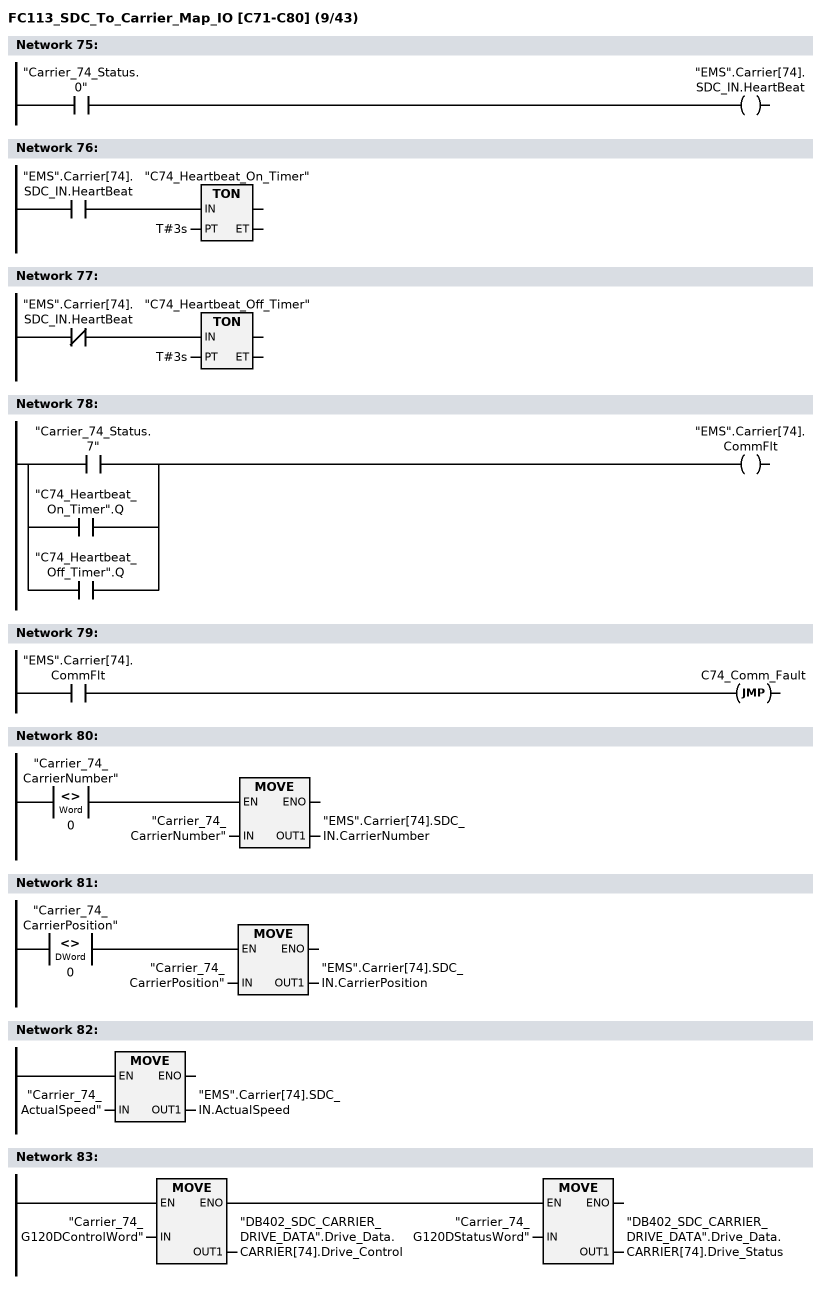
   RUNG wire#powerrail
      Contact( "Carrier_74_Status.0" )
      Coil( "EMS".Carrier[74].SDC_IN.HeartBeat )
   END_RUNG
   // the same network as SCL:
   "EMS".Carrier[74].SDC_IN.HeartBeat := "Carrier_74_Status.0";
END_REGION

REGION Network 76
   "C74_Heartbeat_On_Timer".TON(IN := "EMS".Carrier[74].SDC_IN.HeartBeat, PT := T#3s);
END_REGION

REGION Network 77
   "C74_Heartbeat_Off_Timer".TON(IN := NOT "EMS".Carrier[74].SDC_IN.HeartBeat, PT := T#3s);
END_REGION

REGION Network 78
   RUNG wire#powerrail
      Contact( "Carrier_74_Status.7" )
      wire#w1
      Coil( "EMS".Carrier[74].CommFlt )
   END_RUNG
   RUNG wire#powerrail
      Contact( "C74_Heartbeat_On_Timer".Q )
   END_RUNG wire#w1
   RUNG wire#powerrail
      Contact( "C74_Heartbeat_Off_Timer".Q )
   END_RUNG wire#w1
   // the same network as SCL:
   "EMS".Carrier[74].CommFlt := "Carrier_74_Status.7" OR "C74_Heartbeat_On_Timer".Q OR "C74_Heartbeat_Off_Timer".Q;
END_REGION

REGION Network 79
   RUNG wire#powerrail
      Contact( "EMS".Carrier[74].CommFlt )
      JumpCoil( C74_Comm_Fault )
   END_RUNG
   // the same network as SCL:
   IF "EMS".Carrier[74].CommFlt THEN GOTO C74_Comm_Fault; END_IF;
END_REGION

REGION Network 80
   RUNG wire#powerrail
      { S7_Templates := "SrcType := Word" } NE_Contact(in1 := "Carrier_74_CarrierNumber", in2 := 0)
      Move(in := "Carrier_74_CarrierNumber", out1 => "EMS".Carrier[74].SDC_IN.CarrierNumber)
   END_RUNG
   // the same network as SCL:
   IF "Carrier_74_CarrierNumber" <> 0 THEN
       "EMS".Carrier[74].SDC_IN.CarrierNumber := "Carrier_74_CarrierNumber";
   END_IF;
END_REGION

REGION Network 81
   RUNG wire#powerrail
      { S7_Templates := "SrcType := DWord" } NE_Contact(in1 := "Carrier_74_CarrierPosition", in2 := 0)
      Move(in := "Carrier_74_CarrierPosition", out1 => "EMS".Carrier[74].SDC_IN.CarrierPosition)
   END_RUNG
   // the same network as SCL:
   IF "Carrier_74_CarrierPosition" <> 0 THEN
       "EMS".Carrier[74].SDC_IN.CarrierPosition := "Carrier_74_CarrierPosition";
   END_IF;
END_REGION

REGION Network 82
   RUNG wire#powerrail
      Move(in := "Carrier_74_ActualSpeed", out1 => "EMS".Carrier[74].SDC_IN.ActualSpeed)
   END_RUNG
   // the same network as SCL:
   "EMS".Carrier[74].SDC_IN.ActualSpeed := "Carrier_74_ActualSpeed";
END_REGION

REGION Network 83
   RUNG wire#powerrail
      Move(in := "Carrier_74_G120DControlWord", out1 => "DB402_SDC_CARRIER_DRIVE_DATA".Drive_Data.CARRIER[74].Drive_Control)
      Move(in := "Carrier_74_G120DStatusWord", out1 => "DB402_SDC_CARRIER_DRIVE_DATA".Drive_Data.CARRIER[74].Drive_Status)
   END_RUNG
   // the same network as SCL:
   "DB402_SDC_CARRIER_DRIVE_DATA".Drive_Data.CARRIER[74].Drive_Control := "Carrier_74_G120DControlWord";
   "DB402_SDC_CARRIER_DRIVE_DATA".Drive_Data.CARRIER[74].Drive_Status := "Carrier_74_G120DStatusWord";
END_REGION

REGION Network 84
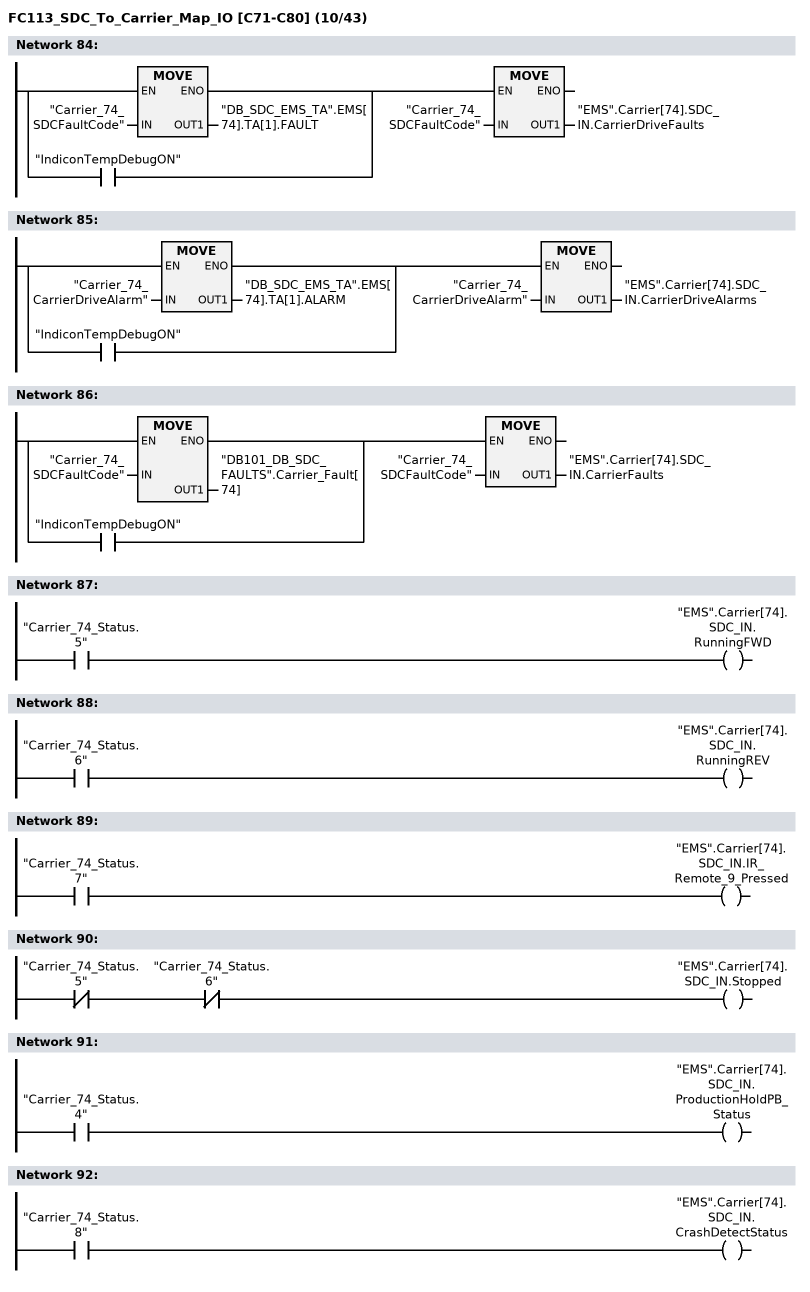
   RUNG wire#powerrail
      Move(in := "Carrier_74_SDCFaultCode", out1 => "DB_SDC_EMS_TA".EMS[74].TA[1].FAULT)
      wire#w1
      Move(in := "Carrier_74_SDCFaultCode", out1 => "EMS".Carrier[74].SDC_IN.CarrierDriveFaults)
   END_RUNG
   RUNG wire#powerrail
      Contact( "IndiconTempDebugON" )
   END_RUNG wire#w1
   // the same network as SCL:
   "DB_SDC_EMS_TA".EMS[74].TA[1].FAULT := "Carrier_74_SDCFaultCode";
   IF TRUE OR "IndiconTempDebugON" THEN
       "EMS".Carrier[74].SDC_IN.CarrierDriveFaults := "Carrier_74_SDCFaultCode";
   END_IF;
END_REGION

REGION Network 85
   RUNG wire#powerrail
      Move(in := "Carrier_74_CarrierDriveAlarm", out1 => "DB_SDC_EMS_TA".EMS[74].TA[1].ALARM)
      wire#w1
      Move(in := "Carrier_74_CarrierDriveAlarm", out1 => "EMS".Carrier[74].SDC_IN.CarrierDriveAlarms)
   END_RUNG
   RUNG wire#powerrail
      Contact( "IndiconTempDebugON" )
   END_RUNG wire#w1
   // the same network as SCL:
   "DB_SDC_EMS_TA".EMS[74].TA[1].ALARM := "Carrier_74_CarrierDriveAlarm";
   IF TRUE OR "IndiconTempDebugON" THEN
       "EMS".Carrier[74].SDC_IN.CarrierDriveAlarms := "Carrier_74_CarrierDriveAlarm";
   END_IF;
END_REGION

REGION Network 86
   RUNG wire#powerrail
      Move(in := "Carrier_74_SDCFaultCode", out1 => "DB101_DB_SDC_FAULTS".Carrier_Fault[74])
      wire#w1
      Move(in := "Carrier_74_SDCFaultCode", out1 => "EMS".Carrier[74].SDC_IN.CarrierFaults)
   END_RUNG
   RUNG wire#powerrail
      Contact( "IndiconTempDebugON" )
   END_RUNG wire#w1
   // the same network as SCL:
   "DB101_DB_SDC_FAULTS".Carrier_Fault[74] := "Carrier_74_SDCFaultCode";
   IF TRUE OR "IndiconTempDebugON" THEN
       "EMS".Carrier[74].SDC_IN.CarrierFaults := "Carrier_74_SDCFaultCode";
   END_IF;
END_REGION

REGION Network 87
   RUNG wire#powerrail
      Contact( "Carrier_74_Status.5" )
      Coil( "EMS".Carrier[74].SDC_IN.RunningFWD )
   END_RUNG
   // the same network as SCL:
   "EMS".Carrier[74].SDC_IN.RunningFWD := "Carrier_74_Status.5";
END_REGION

REGION Network 88
   RUNG wire#powerrail
      Contact( "Carrier_74_Status.6" )
      Coil( "EMS".Carrier[74].SDC_IN.RunningREV )
   END_RUNG
   // the same network as SCL:
   "EMS".Carrier[74].SDC_IN.RunningREV := "Carrier_74_Status.6";
END_REGION

REGION Network 89
   RUNG wire#powerrail
      Contact( "Carrier_74_Status.7" )
      Coil( "EMS".Carrier[74].SDC_IN.IR_Remote_9_Pressed )
   END_RUNG
   // the same network as SCL:
   "EMS".Carrier[74].SDC_IN.IR_Remote_9_Pressed := "Carrier_74_Status.7";
END_REGION

REGION Network 90
   RUNG wire#powerrail
      I_Contact( "Carrier_74_Status.5" )
      I_Contact( "Carrier_74_Status.6" )
      Coil( "EMS".Carrier[74].SDC_IN.Stopped )
   END_RUNG
   // the same network as SCL:
   "EMS".Carrier[74].SDC_IN.Stopped := NOT "Carrier_74_Status.5" AND NOT "Carrier_74_Status.6";
END_REGION

REGION Network 91
   RUNG wire#powerrail
      Contact( "Carrier_74_Status.4" )
      Coil( "EMS".Carrier[74].SDC_IN.ProductionHoldPB_Status )
   END_RUNG
   // the same network as SCL:
   "EMS".Carrier[74].SDC_IN.ProductionHoldPB_Status := "Carrier_74_Status.4";
END_REGION

REGION Network 92
   RUNG wire#powerrail
      Contact( "Carrier_74_Status.8" )
      Coil( "EMS".Carrier[74].SDC_IN.CrashDetectStatus )
   END_RUNG
   // the same network as SCL:
   "EMS".Carrier[74].SDC_IN.CrashDetectStatus := "Carrier_74_Status.8";
END_REGION

REGION Network 93
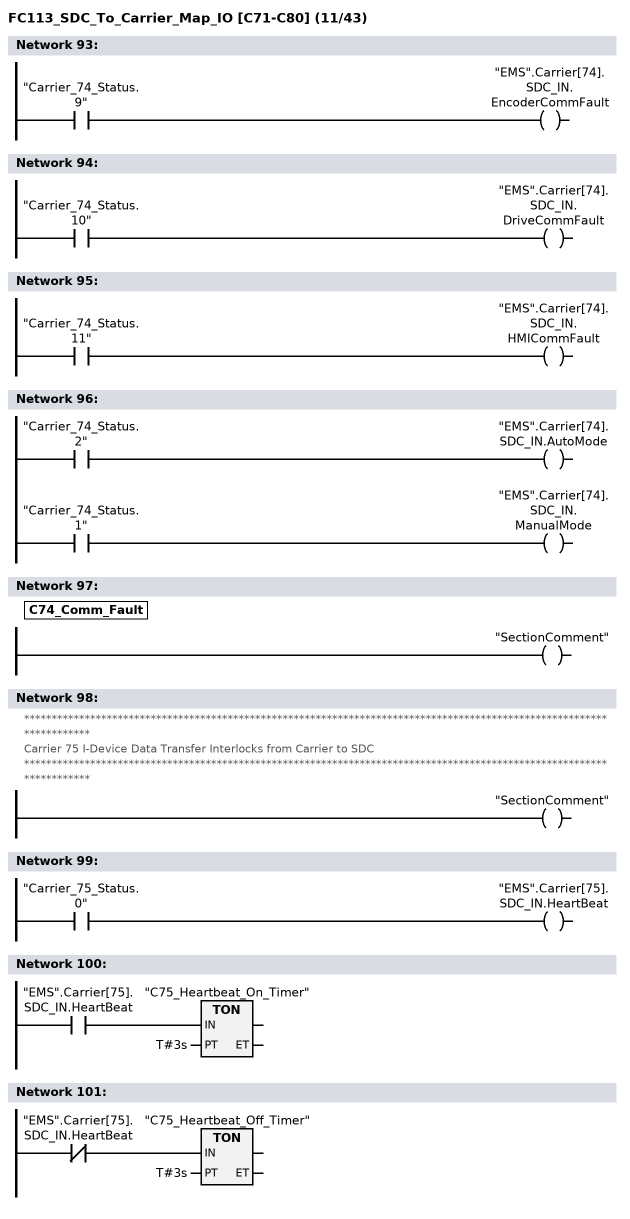
   RUNG wire#powerrail
      Contact( "Carrier_74_Status.9" )
      Coil( "EMS".Carrier[74].SDC_IN.EncoderCommFault )
   END_RUNG
   // the same network as SCL:
   "EMS".Carrier[74].SDC_IN.EncoderCommFault := "Carrier_74_Status.9";
END_REGION

REGION Network 94
   RUNG wire#powerrail
      Contact( "Carrier_74_Status.10" )
      Coil( "EMS".Carrier[74].SDC_IN.DriveCommFault )
   END_RUNG
   // the same network as SCL:
   "EMS".Carrier[74].SDC_IN.DriveCommFault := "Carrier_74_Status.10";
END_REGION

REGION Network 95
   RUNG wire#powerrail
      Contact( "Carrier_74_Status.11" )
      Coil( "EMS".Carrier[74].SDC_IN.HMICommFault )
   END_RUNG
   // the same network as SCL:
   "EMS".Carrier[74].SDC_IN.HMICommFault := "Carrier_74_Status.11";
END_REGION

REGION Network 96
   RUNG wire#powerrail
      Contact( "Carrier_74_Status.2" )
      Coil( "EMS".Carrier[74].SDC_IN.AutoMode )
   END_RUNG
   RUNG wire#powerrail
      Contact( "Carrier_74_Status.1" )
      Coil( "EMS".Carrier[74].SDC_IN.ManualMode )
   END_RUNG
   // the same network as SCL:
   "EMS".Carrier[74].SDC_IN.AutoMode := "Carrier_74_Status.2";
   "EMS".Carrier[74].SDC_IN.ManualMode := "Carrier_74_Status.1";
END_REGION

REGION Network 97
   Label( C74_Comm_Fault )
   RUNG wire#powerrail
      Coil( "SectionComment" )
   END_RUNG
   // the same network as SCL:
   C74_Comm_Fault:
   "SectionComment" := TRUE;
END_REGION

REGION Network 98
   // **********************************************************************************************************************
   // 
   // Carrier 75 I-Device Data Transfer Interlocks from Carrier to SDC
   // 
   // **********************************************************************************************************************
   RUNG wire#powerrail
      Coil( "SectionComment" )
   END_RUNG
   // the same network as SCL:
   "SectionComment" := TRUE;
END_REGION

REGION Network 99
   RUNG wire#powerrail
      Contact( "Carrier_75_Status.0" )
      Coil( "EMS".Carrier[75].SDC_IN.HeartBeat )
   END_RUNG
   // the same network as SCL:
   "EMS".Carrier[75].SDC_IN.HeartBeat := "Carrier_75_Status.0";
END_REGION

REGION Network 100
   "C75_Heartbeat_On_Timer".TON(IN := "EMS".Carrier[75].SDC_IN.HeartBeat, PT := T#3s);
END_REGION

REGION Network 101
   "C75_Heartbeat_Off_Timer".TON(IN := NOT "EMS".Carrier[75].SDC_IN.HeartBeat, PT := T#3s);
END_REGION

REGION Network 102
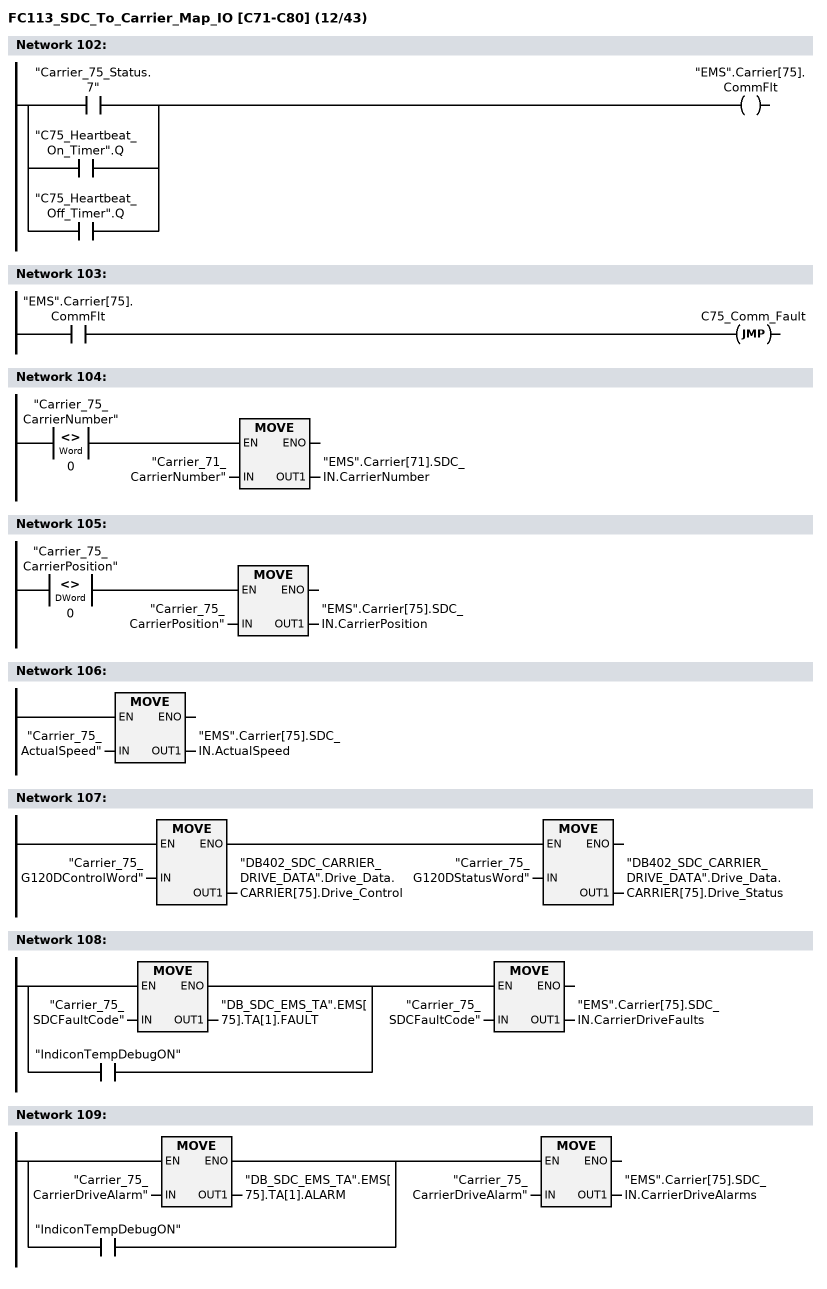
   RUNG wire#powerrail
      Contact( "Carrier_75_Status.7" )
      wire#w1
      Coil( "EMS".Carrier[75].CommFlt )
   END_RUNG
   RUNG wire#powerrail
      Contact( "C75_Heartbeat_On_Timer".Q )
   END_RUNG wire#w1
   RUNG wire#powerrail
      Contact( "C75_Heartbeat_Off_Timer".Q )
   END_RUNG wire#w1
   // the same network as SCL:
   "EMS".Carrier[75].CommFlt := "Carrier_75_Status.7" OR "C75_Heartbeat_On_Timer".Q OR "C75_Heartbeat_Off_Timer".Q;
END_REGION

REGION Network 103
   RUNG wire#powerrail
      Contact( "EMS".Carrier[75].CommFlt )
      JumpCoil( C75_Comm_Fault )
   END_RUNG
   // the same network as SCL:
   IF "EMS".Carrier[75].CommFlt THEN GOTO C75_Comm_Fault; END_IF;
END_REGION

REGION Network 104
   RUNG wire#powerrail
      { S7_Templates := "SrcType := Word" } NE_Contact(in1 := "Carrier_75_CarrierNumber", in2 := 0)
      Move(in := "Carrier_71_CarrierNumber", out1 => "EMS".Carrier[71].SDC_IN.CarrierNumber)
   END_RUNG
   // the same network as SCL:
   IF "Carrier_75_CarrierNumber" <> 0 THEN
       "EMS".Carrier[71].SDC_IN.CarrierNumber := "Carrier_71_CarrierNumber";
   END_IF;
END_REGION

REGION Network 105
   RUNG wire#powerrail
      { S7_Templates := "SrcType := DWord" } NE_Contact(in1 := "Carrier_75_CarrierPosition", in2 := 0)
      Move(in := "Carrier_75_CarrierPosition", out1 => "EMS".Carrier[75].SDC_IN.CarrierPosition)
   END_RUNG
   // the same network as SCL:
   IF "Carrier_75_CarrierPosition" <> 0 THEN
       "EMS".Carrier[75].SDC_IN.CarrierPosition := "Carrier_75_CarrierPosition";
   END_IF;
END_REGION

REGION Network 106
   RUNG wire#powerrail
      Move(in := "Carrier_75_ActualSpeed", out1 => "EMS".Carrier[75].SDC_IN.ActualSpeed)
   END_RUNG
   // the same network as SCL:
   "EMS".Carrier[75].SDC_IN.ActualSpeed := "Carrier_75_ActualSpeed";
END_REGION

REGION Network 107
   RUNG wire#powerrail
      Move(in := "Carrier_75_G120DControlWord", out1 => "DB402_SDC_CARRIER_DRIVE_DATA".Drive_Data.CARRIER[75].Drive_Control)
      Move(in := "Carrier_75_G120DStatusWord", out1 => "DB402_SDC_CARRIER_DRIVE_DATA".Drive_Data.CARRIER[75].Drive_Status)
   END_RUNG
   // the same network as SCL:
   "DB402_SDC_CARRIER_DRIVE_DATA".Drive_Data.CARRIER[75].Drive_Control := "Carrier_75_G120DControlWord";
   "DB402_SDC_CARRIER_DRIVE_DATA".Drive_Data.CARRIER[75].Drive_Status := "Carrier_75_G120DStatusWord";
END_REGION

REGION Network 108
   RUNG wire#powerrail
      Move(in := "Carrier_75_SDCFaultCode", out1 => "DB_SDC_EMS_TA".EMS[75].TA[1].FAULT)
      wire#w1
      Move(in := "Carrier_75_SDCFaultCode", out1 => "EMS".Carrier[75].SDC_IN.CarrierDriveFaults)
   END_RUNG
   RUNG wire#powerrail
      Contact( "IndiconTempDebugON" )
   END_RUNG wire#w1
   // the same network as SCL:
   "DB_SDC_EMS_TA".EMS[75].TA[1].FAULT := "Carrier_75_SDCFaultCode";
   IF TRUE OR "IndiconTempDebugON" THEN
       "EMS".Carrier[75].SDC_IN.CarrierDriveFaults := "Carrier_75_SDCFaultCode";
   END_IF;
END_REGION

REGION Network 109
   RUNG wire#powerrail
      Move(in := "Carrier_75_CarrierDriveAlarm", out1 => "DB_SDC_EMS_TA".EMS[75].TA[1].ALARM)
      wire#w1
      Move(in := "Carrier_75_CarrierDriveAlarm", out1 => "EMS".Carrier[75].SDC_IN.CarrierDriveAlarms)
   END_RUNG
   RUNG wire#powerrail
      Contact( "IndiconTempDebugON" )
   END_RUNG wire#w1
   // the same network as SCL:
   "DB_SDC_EMS_TA".EMS[75].TA[1].ALARM := "Carrier_75_CarrierDriveAlarm";
   IF TRUE OR "IndiconTempDebugON" THEN
       "EMS".Carrier[75].SDC_IN.CarrierDriveAlarms := "Carrier_75_CarrierDriveAlarm";
   END_IF;
END_REGION

REGION Network 110
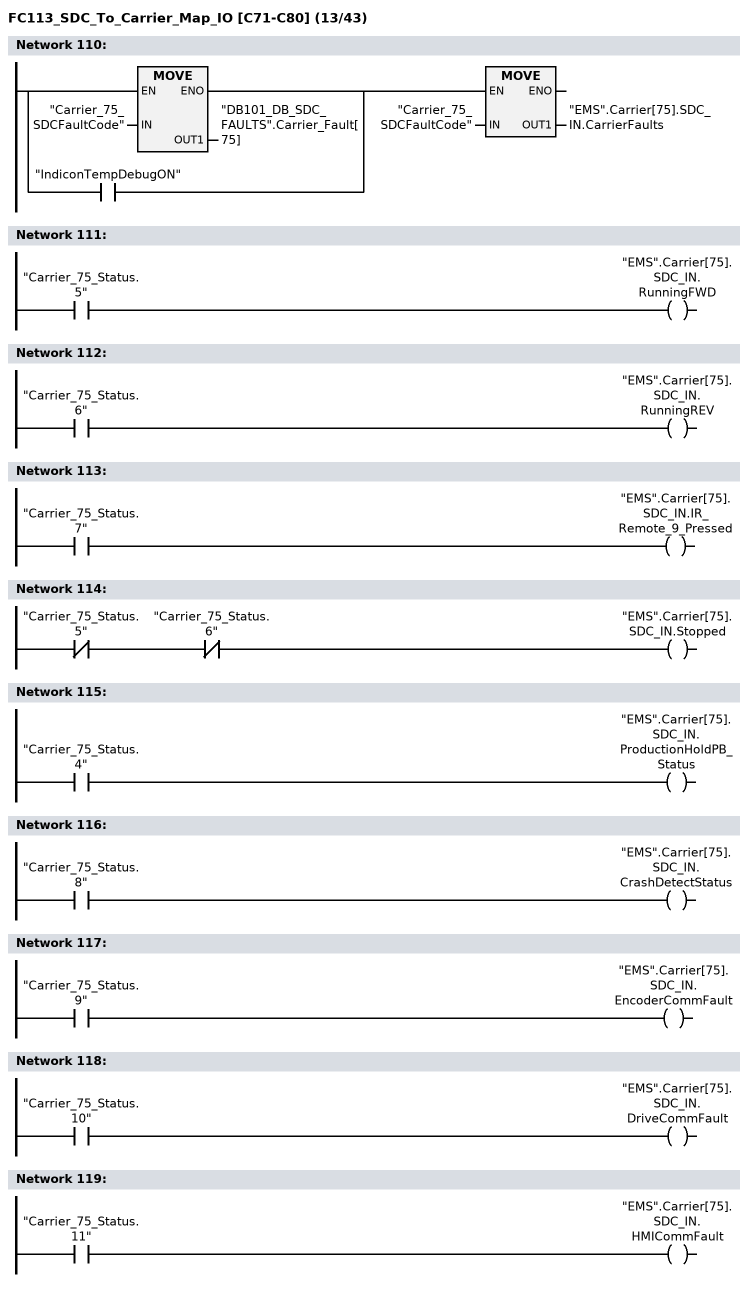
   RUNG wire#powerrail
      Move(in := "Carrier_75_SDCFaultCode", out1 => "DB101_DB_SDC_FAULTS".Carrier_Fault[75])
      wire#w1
      Move(in := "Carrier_75_SDCFaultCode", out1 => "EMS".Carrier[75].SDC_IN.CarrierFaults)
   END_RUNG
   RUNG wire#powerrail
      Contact( "IndiconTempDebugON" )
   END_RUNG wire#w1
   // the same network as SCL:
   "DB101_DB_SDC_FAULTS".Carrier_Fault[75] := "Carrier_75_SDCFaultCode";
   IF TRUE OR "IndiconTempDebugON" THEN
       "EMS".Carrier[75].SDC_IN.CarrierFaults := "Carrier_75_SDCFaultCode";
   END_IF;
END_REGION

REGION Network 111
   RUNG wire#powerrail
      Contact( "Carrier_75_Status.5" )
      Coil( "EMS".Carrier[75].SDC_IN.RunningFWD )
   END_RUNG
   // the same network as SCL:
   "EMS".Carrier[75].SDC_IN.RunningFWD := "Carrier_75_Status.5";
END_REGION

REGION Network 112
   RUNG wire#powerrail
      Contact( "Carrier_75_Status.6" )
      Coil( "EMS".Carrier[75].SDC_IN.RunningREV )
   END_RUNG
   // the same network as SCL:
   "EMS".Carrier[75].SDC_IN.RunningREV := "Carrier_75_Status.6";
END_REGION

REGION Network 113
   RUNG wire#powerrail
      Contact( "Carrier_75_Status.7" )
      Coil( "EMS".Carrier[75].SDC_IN.IR_Remote_9_Pressed )
   END_RUNG
   // the same network as SCL:
   "EMS".Carrier[75].SDC_IN.IR_Remote_9_Pressed := "Carrier_75_Status.7";
END_REGION

REGION Network 114
   RUNG wire#powerrail
      I_Contact( "Carrier_75_Status.5" )
      I_Contact( "Carrier_75_Status.6" )
      Coil( "EMS".Carrier[75].SDC_IN.Stopped )
   END_RUNG
   // the same network as SCL:
   "EMS".Carrier[75].SDC_IN.Stopped := NOT "Carrier_75_Status.5" AND NOT "Carrier_75_Status.6";
END_REGION

REGION Network 115
   RUNG wire#powerrail
      Contact( "Carrier_75_Status.4" )
      Coil( "EMS".Carrier[75].SDC_IN.ProductionHoldPB_Status )
   END_RUNG
   // the same network as SCL:
   "EMS".Carrier[75].SDC_IN.ProductionHoldPB_Status := "Carrier_75_Status.4";
END_REGION

REGION Network 116
   RUNG wire#powerrail
      Contact( "Carrier_75_Status.8" )
      Coil( "EMS".Carrier[75].SDC_IN.CrashDetectStatus )
   END_RUNG
   // the same network as SCL:
   "EMS".Carrier[75].SDC_IN.CrashDetectStatus := "Carrier_75_Status.8";
END_REGION

REGION Network 117
   RUNG wire#powerrail
      Contact( "Carrier_75_Status.9" )
      Coil( "EMS".Carrier[75].SDC_IN.EncoderCommFault )
   END_RUNG
   // the same network as SCL:
   "EMS".Carrier[75].SDC_IN.EncoderCommFault := "Carrier_75_Status.9";
END_REGION

REGION Network 118
   RUNG wire#powerrail
      Contact( "Carrier_75_Status.10" )
      Coil( "EMS".Carrier[75].SDC_IN.DriveCommFault )
   END_RUNG
   // the same network as SCL:
   "EMS".Carrier[75].SDC_IN.DriveCommFault := "Carrier_75_Status.10";
END_REGION

REGION Network 119
   RUNG wire#powerrail
      Contact( "Carrier_75_Status.11" )
      Coil( "EMS".Carrier[75].SDC_IN.HMICommFault )
   END_RUNG
   // the same network as SCL:
   "EMS".Carrier[75].SDC_IN.HMICommFault := "Carrier_75_Status.11";
END_REGION

REGION Network 120
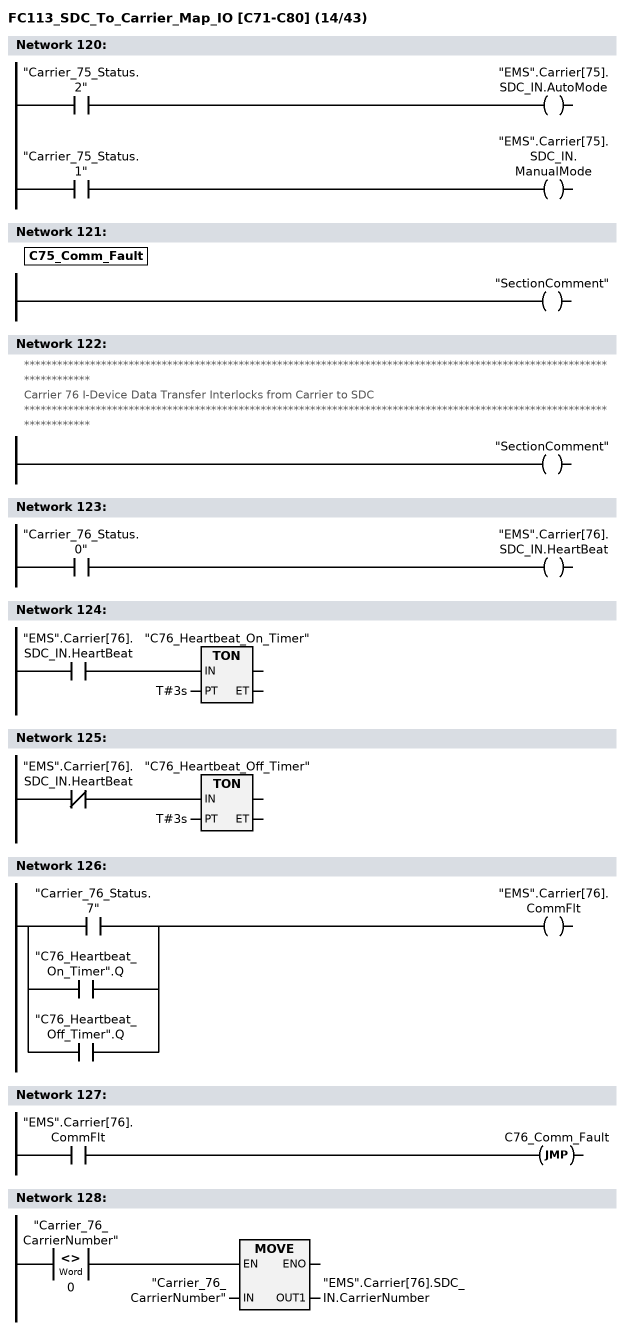
   RUNG wire#powerrail
      Contact( "Carrier_75_Status.2" )
      Coil( "EMS".Carrier[75].SDC_IN.AutoMode )
   END_RUNG
   RUNG wire#powerrail
      Contact( "Carrier_75_Status.1" )
      Coil( "EMS".Carrier[75].SDC_IN.ManualMode )
   END_RUNG
   // the same network as SCL:
   "EMS".Carrier[75].SDC_IN.AutoMode := "Carrier_75_Status.2";
   "EMS".Carrier[75].SDC_IN.ManualMode := "Carrier_75_Status.1";
END_REGION

REGION Network 121
   Label( C75_Comm_Fault )
   RUNG wire#powerrail
      Coil( "SectionComment" )
   END_RUNG
   // the same network as SCL:
   C75_Comm_Fault:
   "SectionComment" := TRUE;
END_REGION

REGION Network 122
   // **********************************************************************************************************************
   // 
   // Carrier 76 I-Device Data Transfer Interlocks from Carrier to SDC
   // 
   // **********************************************************************************************************************
   RUNG wire#powerrail
      Coil( "SectionComment" )
   END_RUNG
   // the same network as SCL:
   "SectionComment" := TRUE;
END_REGION

REGION Network 123
   RUNG wire#powerrail
      Contact( "Carrier_76_Status.0" )
      Coil( "EMS".Carrier[76].SDC_IN.HeartBeat )
   END_RUNG
   // the same network as SCL:
   "EMS".Carrier[76].SDC_IN.HeartBeat := "Carrier_76_Status.0";
END_REGION

REGION Network 124
   "C76_Heartbeat_On_Timer".TON(IN := "EMS".Carrier[76].SDC_IN.HeartBeat, PT := T#3s);
END_REGION

REGION Network 125
   "C76_Heartbeat_Off_Timer".TON(IN := NOT "EMS".Carrier[76].SDC_IN.HeartBeat, PT := T#3s);
END_REGION

REGION Network 126
   RUNG wire#powerrail
      Contact( "Carrier_76_Status.7" )
      wire#w1
      Coil( "EMS".Carrier[76].CommFlt )
   END_RUNG
   RUNG wire#powerrail
      Contact( "C76_Heartbeat_On_Timer".Q )
   END_RUNG wire#w1
   RUNG wire#powerrail
      Contact( "C76_Heartbeat_Off_Timer".Q )
   END_RUNG wire#w1
   // the same network as SCL:
   "EMS".Carrier[76].CommFlt := "Carrier_76_Status.7" OR "C76_Heartbeat_On_Timer".Q OR "C76_Heartbeat_Off_Timer".Q;
END_REGION

REGION Network 127
   RUNG wire#powerrail
      Contact( "EMS".Carrier[76].CommFlt )
      JumpCoil( C76_Comm_Fault )
   END_RUNG
   // the same network as SCL:
   IF "EMS".Carrier[76].CommFlt THEN GOTO C76_Comm_Fault; END_IF;
END_REGION

REGION Network 128
   RUNG wire#powerrail
      { S7_Templates := "SrcType := Word" } NE_Contact(in1 := "Carrier_76_CarrierNumber", in2 := 0)
      Move(in := "Carrier_76_CarrierNumber", out1 => "EMS".Carrier[76].SDC_IN.CarrierNumber)
   END_RUNG
   // the same network as SCL:
   IF "Carrier_76_CarrierNumber" <> 0 THEN
       "EMS".Carrier[76].SDC_IN.CarrierNumber := "Carrier_76_CarrierNumber";
   END_IF;
END_REGION

REGION Network 129
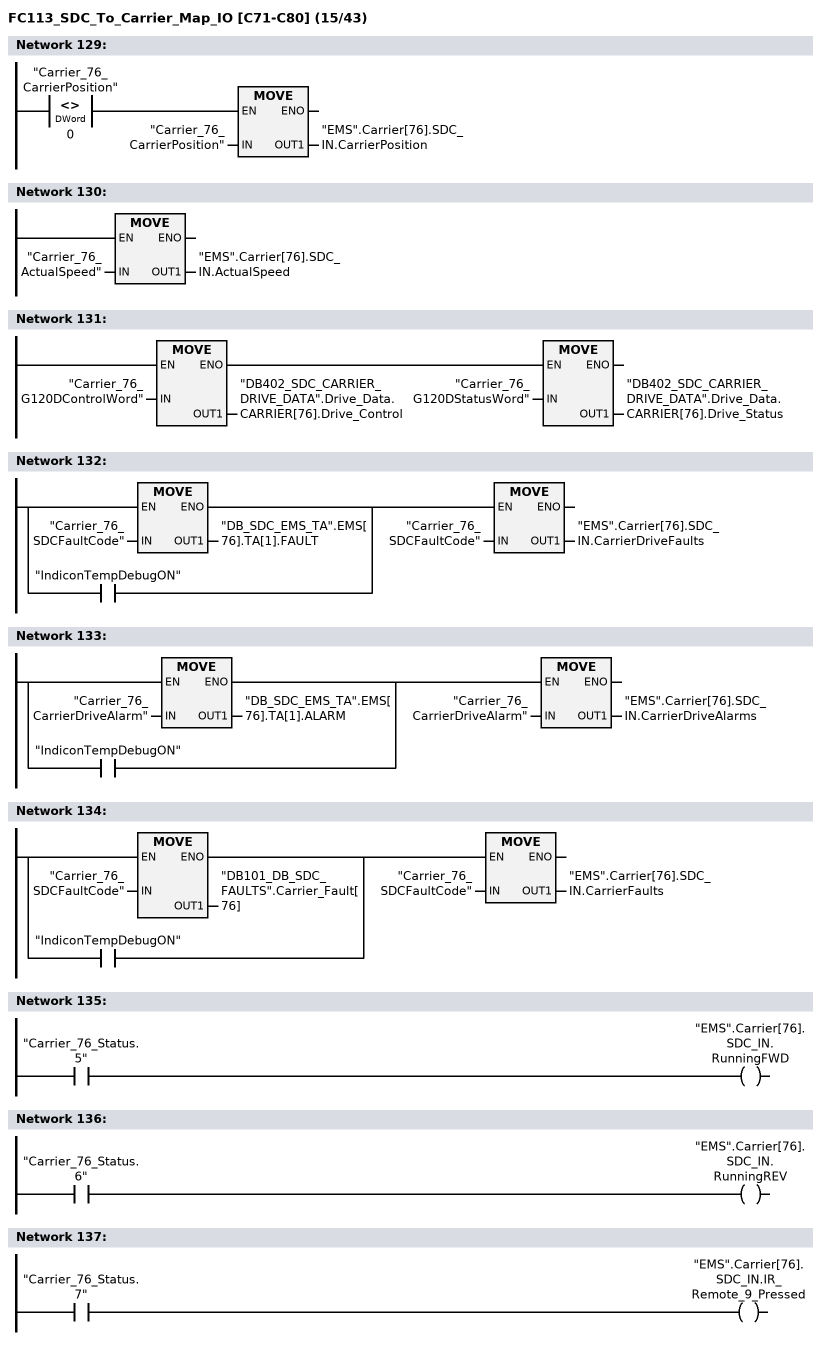
   RUNG wire#powerrail
      { S7_Templates := "SrcType := DWord" } NE_Contact(in1 := "Carrier_76_CarrierPosition", in2 := 0)
      Move(in := "Carrier_76_CarrierPosition", out1 => "EMS".Carrier[76].SDC_IN.CarrierPosition)
   END_RUNG
   // the same network as SCL:
   IF "Carrier_76_CarrierPosition" <> 0 THEN
       "EMS".Carrier[76].SDC_IN.CarrierPosition := "Carrier_76_CarrierPosition";
   END_IF;
END_REGION

REGION Network 130
   RUNG wire#powerrail
      Move(in := "Carrier_76_ActualSpeed", out1 => "EMS".Carrier[76].SDC_IN.ActualSpeed)
   END_RUNG
   // the same network as SCL:
   "EMS".Carrier[76].SDC_IN.ActualSpeed := "Carrier_76_ActualSpeed";
END_REGION

REGION Network 131
   RUNG wire#powerrail
      Move(in := "Carrier_76_G120DControlWord", out1 => "DB402_SDC_CARRIER_DRIVE_DATA".Drive_Data.CARRIER[76].Drive_Control)
      Move(in := "Carrier_76_G120DStatusWord", out1 => "DB402_SDC_CARRIER_DRIVE_DATA".Drive_Data.CARRIER[76].Drive_Status)
   END_RUNG
   // the same network as SCL:
   "DB402_SDC_CARRIER_DRIVE_DATA".Drive_Data.CARRIER[76].Drive_Control := "Carrier_76_G120DControlWord";
   "DB402_SDC_CARRIER_DRIVE_DATA".Drive_Data.CARRIER[76].Drive_Status := "Carrier_76_G120DStatusWord";
END_REGION

REGION Network 132
   RUNG wire#powerrail
      Move(in := "Carrier_76_SDCFaultCode", out1 => "DB_SDC_EMS_TA".EMS[76].TA[1].FAULT)
      wire#w1
      Move(in := "Carrier_76_SDCFaultCode", out1 => "EMS".Carrier[76].SDC_IN.CarrierDriveFaults)
   END_RUNG
   RUNG wire#powerrail
      Contact( "IndiconTempDebugON" )
   END_RUNG wire#w1
   // the same network as SCL:
   "DB_SDC_EMS_TA".EMS[76].TA[1].FAULT := "Carrier_76_SDCFaultCode";
   IF TRUE OR "IndiconTempDebugON" THEN
       "EMS".Carrier[76].SDC_IN.CarrierDriveFaults := "Carrier_76_SDCFaultCode";
   END_IF;
END_REGION

REGION Network 133
   RUNG wire#powerrail
      Move(in := "Carrier_76_CarrierDriveAlarm", out1 => "DB_SDC_EMS_TA".EMS[76].TA[1].ALARM)
      wire#w1
      Move(in := "Carrier_76_CarrierDriveAlarm", out1 => "EMS".Carrier[76].SDC_IN.CarrierDriveAlarms)
   END_RUNG
   RUNG wire#powerrail
      Contact( "IndiconTempDebugON" )
   END_RUNG wire#w1
   // the same network as SCL:
   "DB_SDC_EMS_TA".EMS[76].TA[1].ALARM := "Carrier_76_CarrierDriveAlarm";
   IF TRUE OR "IndiconTempDebugON" THEN
       "EMS".Carrier[76].SDC_IN.CarrierDriveAlarms := "Carrier_76_CarrierDriveAlarm";
   END_IF;
END_REGION

REGION Network 134
   RUNG wire#powerrail
      Move(in := "Carrier_76_SDCFaultCode", out1 => "DB101_DB_SDC_FAULTS".Carrier_Fault[76])
      wire#w1
      Move(in := "Carrier_76_SDCFaultCode", out1 => "EMS".Carrier[76].SDC_IN.CarrierFaults)
   END_RUNG
   RUNG wire#powerrail
      Contact( "IndiconTempDebugON" )
   END_RUNG wire#w1
   // the same network as SCL:
   "DB101_DB_SDC_FAULTS".Carrier_Fault[76] := "Carrier_76_SDCFaultCode";
   IF TRUE OR "IndiconTempDebugON" THEN
       "EMS".Carrier[76].SDC_IN.CarrierFaults := "Carrier_76_SDCFaultCode";
   END_IF;
END_REGION

REGION Network 135
   RUNG wire#powerrail
      Contact( "Carrier_76_Status.5" )
      Coil( "EMS".Carrier[76].SDC_IN.RunningFWD )
   END_RUNG
   // the same network as SCL:
   "EMS".Carrier[76].SDC_IN.RunningFWD := "Carrier_76_Status.5";
END_REGION

REGION Network 136
   RUNG wire#powerrail
      Contact( "Carrier_76_Status.6" )
      Coil( "EMS".Carrier[76].SDC_IN.RunningREV )
   END_RUNG
   // the same network as SCL:
   "EMS".Carrier[76].SDC_IN.RunningREV := "Carrier_76_Status.6";
END_REGION

REGION Network 137
   RUNG wire#powerrail
      Contact( "Carrier_76_Status.7" )
      Coil( "EMS".Carrier[76].SDC_IN.IR_Remote_9_Pressed )
   END_RUNG
   // the same network as SCL:
   "EMS".Carrier[76].SDC_IN.IR_Remote_9_Pressed := "Carrier_76_Status.7";
END_REGION

REGION Network 138
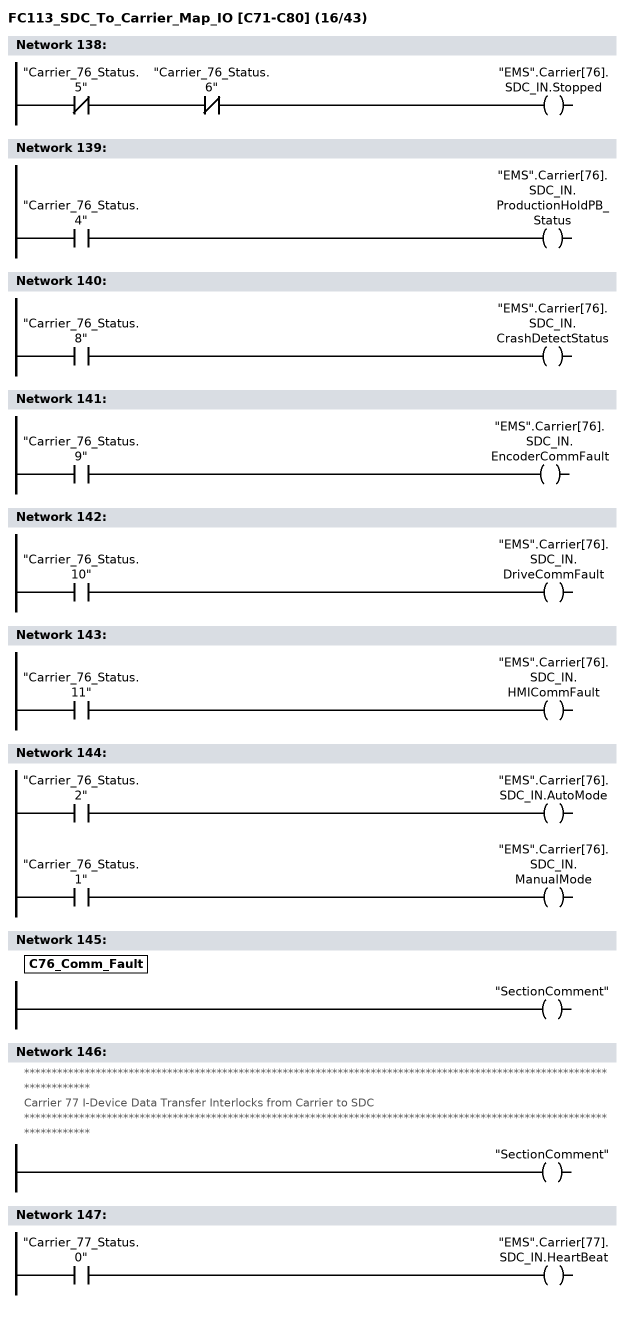
   RUNG wire#powerrail
      I_Contact( "Carrier_76_Status.5" )
      I_Contact( "Carrier_76_Status.6" )
      Coil( "EMS".Carrier[76].SDC_IN.Stopped )
   END_RUNG
   // the same network as SCL:
   "EMS".Carrier[76].SDC_IN.Stopped := NOT "Carrier_76_Status.5" AND NOT "Carrier_76_Status.6";
END_REGION

REGION Network 139
   RUNG wire#powerrail
      Contact( "Carrier_76_Status.4" )
      Coil( "EMS".Carrier[76].SDC_IN.ProductionHoldPB_Status )
   END_RUNG
   // the same network as SCL:
   "EMS".Carrier[76].SDC_IN.ProductionHoldPB_Status := "Carrier_76_Status.4";
END_REGION

REGION Network 140
   RUNG wire#powerrail
      Contact( "Carrier_76_Status.8" )
      Coil( "EMS".Carrier[76].SDC_IN.CrashDetectStatus )
   END_RUNG
   // the same network as SCL:
   "EMS".Carrier[76].SDC_IN.CrashDetectStatus := "Carrier_76_Status.8";
END_REGION

REGION Network 141
   RUNG wire#powerrail
      Contact( "Carrier_76_Status.9" )
      Coil( "EMS".Carrier[76].SDC_IN.EncoderCommFault )
   END_RUNG
   // the same network as SCL:
   "EMS".Carrier[76].SDC_IN.EncoderCommFault := "Carrier_76_Status.9";
END_REGION

REGION Network 142
   RUNG wire#powerrail
      Contact( "Carrier_76_Status.10" )
      Coil( "EMS".Carrier[76].SDC_IN.DriveCommFault )
   END_RUNG
   // the same network as SCL:
   "EMS".Carrier[76].SDC_IN.DriveCommFault := "Carrier_76_Status.10";
END_REGION

REGION Network 143
   RUNG wire#powerrail
      Contact( "Carrier_76_Status.11" )
      Coil( "EMS".Carrier[76].SDC_IN.HMICommFault )
   END_RUNG
   // the same network as SCL:
   "EMS".Carrier[76].SDC_IN.HMICommFault := "Carrier_76_Status.11";
END_REGION

REGION Network 144
   RUNG wire#powerrail
      Contact( "Carrier_76_Status.2" )
      Coil( "EMS".Carrier[76].SDC_IN.AutoMode )
   END_RUNG
   RUNG wire#powerrail
      Contact( "Carrier_76_Status.1" )
      Coil( "EMS".Carrier[76].SDC_IN.ManualMode )
   END_RUNG
   // the same network as SCL:
   "EMS".Carrier[76].SDC_IN.AutoMode := "Carrier_76_Status.2";
   "EMS".Carrier[76].SDC_IN.ManualMode := "Carrier_76_Status.1";
END_REGION
